REGION Network 9
   RUNG wire#powerrail
      Contact( "DB120".Static_81 )
      Contact( "TsinReq6" )
      wire#w1
      Coil( "DB127".Static_82 )
   END_RUNG
   RUNG wire#powerrail
      Contact( "DB120".Static_89 )
      Contact( "DB88".Static_8 )
   END_RUNG wire#w1
   // the same network as SCL:
   "DB127".Static_82 := ("DB120".Static_81 AND "TsinReq6") OR ("DB120".Static_89 AND "DB88".Static_8);
END_REGION

REGION Network 10
   RUNG wire#powerrail
      Contact( "DB120".Static_80 )
      I_Contact( "DB121".Static_75 )
      wire#w1
      Contact( "DB88".Static_17 )
      Coil( "DB127".Static_89 )
   END_RUNG
   RUNG wire#powerrail
      Contact( "DB120".Static_88 )
      I_Contact( "DB121".Static_75 )
   END_RUNG wire#w1
   RUNG wire#powerrail
      Contact( "DB120".Static_82 )
      I_Contact( "DB88".Static_8 )
   END_RUNG wire#w1
   // the same network as SCL:
   "DB127".Static_89 := (("DB120".Static_80 AND NOT "DB121".Static_75) OR ("DB120".Static_88 AND NOT "DB121".Static_75) OR ("DB120".Static_82 AND NOT "DB88".Static_8)) AND "DB88".Static_17;
END_REGION

REGION Network 11
   #_w1 := "DB121".Static_75 AND NOT "flReqMch6";   // rising edge
   "flReqMch6" := "DB121".Static_75;
   "DB127".Static_83 := ("DB120".Static_88 AND ("MC006-CO" OR "DB88".Static_8)) OR ("DB120".Static_84 AND NOT "DB121".Static_94 AND NOT "DB88".Static_19) OR ("DB120".Static_82 AND ("DB88".Static_19 OR "DB121".Static_94 OR "DB121".Static_75) AND "DB88".Static_8) OR (#_w1 AND "DB120".Static_82 AND "DB88".Static_8);
END_REGION

REGION Network 12
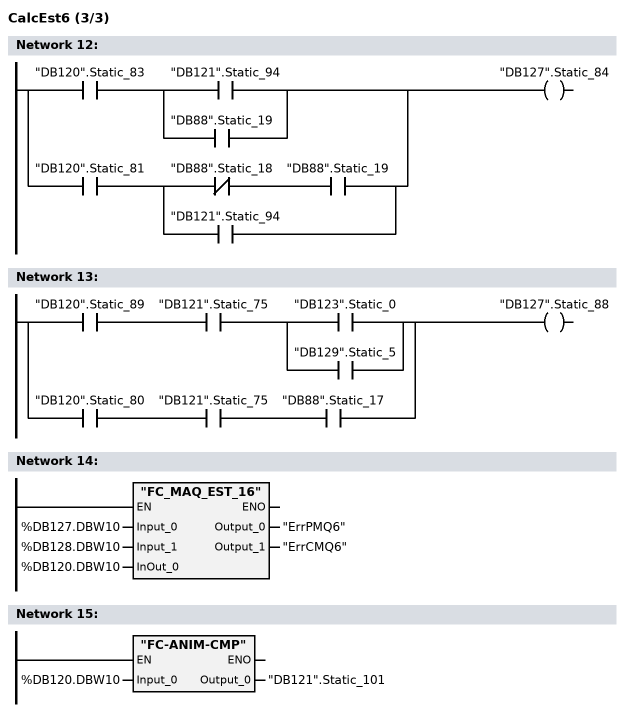
   "DB127".Static_84 := ("DB120".Static_83 AND ("DB121".Static_94 OR "DB88".Static_19)) OR ("DB120".Static_81 AND ("DB121".Static_94 OR (NOT "DB88".Static_18 AND "DB88".Static_19)));
END_REGION

REGION Network 13
   "DB127".Static_88 := ("DB120".Static_89 AND "DB121".Static_75 AND ("DB123".Static_0 OR "DB129".Static_5)) OR ("DB120".Static_80 AND "DB121".Static_75 AND "DB88".Static_17);
END_REGION

REGION Network 14
   RUNG wire#powerrail
      "FC_MAQ_EST_16"(Input_0 := %DB127.DBW10, Input_1 := %DB128.DBW10, Output_0 => "ErrPMQ6", Output_1 => "ErrCMQ6", InOut_0 := %DB120.DBW10)
   END_RUNG
   // the same network as SCL:
   "FC_MAQ_EST_16"(Input_0 := %DB127.DBW10,
                   Input_1 := %DB128.DBW10,
                   InOut_0 := %DB120.DBW10,
                   Output_0 => "ErrPMQ6",
                   Output_1 => "ErrCMQ6");
END_REGION

REGION Network 15
   RUNG wire#powerrail
      "FC-ANIM-CMP"(Input_0 := %DB120.DBW10, Output_0 => "DB121".Static_101)
   END_RUNG
   // the same network as SCL:
   "FC-ANIM-CMP"(Input_0 := %DB120.DBW10, Output_0 => "DB121".Static_101);
END_REGION
END_FUNCTION

// folder: Compresores/Baja

FUNCTION "AutoCmpBaja" : Void   // FC24, LAD
{ S7_Optimized_Access := 'FALSE' }
VERSION : 0.1
   VAR_TEMP   // added for the SCL form of the ladder/FBD networks
      _w1 : Bool;
      _s5time1 : S5Time;
      _w2 : Bool;
   END_VAR
BEGIN

REGION Network 1 (STL)
         A(;
         L     "CmpBajaAuto".Static_10;
         L     "CmpBajaAuto".Static_5;
         <=R;
         );
         JNB   M001;
         L     "CmpBajaAuto".Static_5;
         L     1;
         +R;
         T     "CmpBajaAuto".Static_10;
   M001: NOP   0;
END_REGION

REGION Network 2 (STL)
         A(;
         L     "CmpBajaAuto".Static_11;
         L     "CmpBajaAuto".Static_6;
         <=R;
         );
         JNB   M002;
         L     "CmpBajaAuto".Static_6;
         L     1;
         +R;
         T     "CmpBajaAuto".Static_11;
   M002: NOP   0;
END_REGION

REGION Network 3 (STL)
         A(;
         L     "CmpBajaAuto".Static_12;
         L     "CmpBajaAuto".Static_7;
         <=R;
         );
         JNB   M003;
         L     "CmpBajaAuto".Static_7;
         L     1;
         +R;
         T     "CmpBajaAuto".Static_12;
   M003: NOP   0;
END_REGION

REGION Network 4 (STL)
         A(;
         L     "CmpBajaAuto".Static_13;
         L     "CmpBajaAuto".Static_8;
         <=R;
         );
         JNB   M004;
         L     "CmpBajaAuto".Static_8;
         L     1;
         +R;
         T     "CmpBajaAuto".Static_13;
   M004: NOP   0;
END_REGION

REGION Network 5 (STL)
         A(;
         L     "CmpBajaAuto".Static_14;
         L     "CmpBajaAuto".Static_9;
         <=R;
         );
         JNB   M005;
         L     "CmpBajaAuto".Static_9;
         L     1;
         +R;
         T     "CmpBajaAuto".Static_14;
   M005: NOP   0;
END_REGION

REGION Network 6
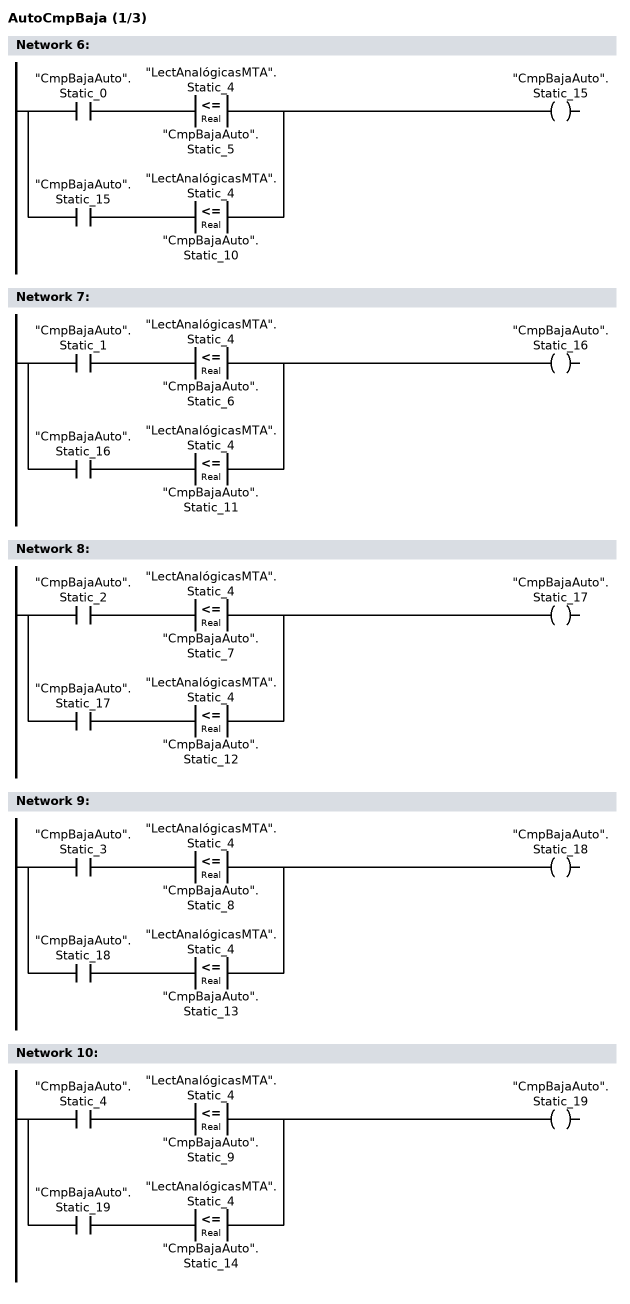
   "CmpBajaAuto".Static_15 := ("CmpBajaAuto".Static_0 AND ("LectAnalógicasMTA".Static_4 <= "CmpBajaAuto".Static_5)) OR ("CmpBajaAuto".Static_15 AND ("LectAnalógicasMTA".Static_4 <= "CmpBajaAuto".Static_10));
END_REGION

REGION Network 7
   "CmpBajaAuto".Static_16 := ("CmpBajaAuto".Static_1 AND ("LectAnalógicasMTA".Static_4 <= "CmpBajaAuto".Static_6)) OR ("CmpBajaAuto".Static_16 AND ("LectAnalógicasMTA".Static_4 <= "CmpBajaAuto".Static_11));
END_REGION

REGION Network 8
   "CmpBajaAuto".Static_17 := ("CmpBajaAuto".Static_2 AND ("LectAnalógicasMTA".Static_4 <= "CmpBajaAuto".Static_7)) OR ("CmpBajaAuto".Static_17 AND ("LectAnalógicasMTA".Static_4 <= "CmpBajaAuto".Static_12));
END_REGION

REGION Network 9
   "CmpBajaAuto".Static_18 := ("CmpBajaAuto".Static_3 AND ("LectAnalógicasMTA".Static_4 <= "CmpBajaAuto".Static_8)) OR ("CmpBajaAuto".Static_18 AND ("LectAnalógicasMTA".Static_4 <= "CmpBajaAuto".Static_13));
END_REGION

REGION Network 10
   "CmpBajaAuto".Static_19 := ("CmpBajaAuto".Static_4 AND ("LectAnalógicasMTA".Static_4 <= "CmpBajaAuto".Static_9)) OR ("CmpBajaAuto".Static_19 AND ("LectAnalógicasMTA".Static_4 <= "CmpBajaAuto".Static_14));
END_REGION

REGION Network 11
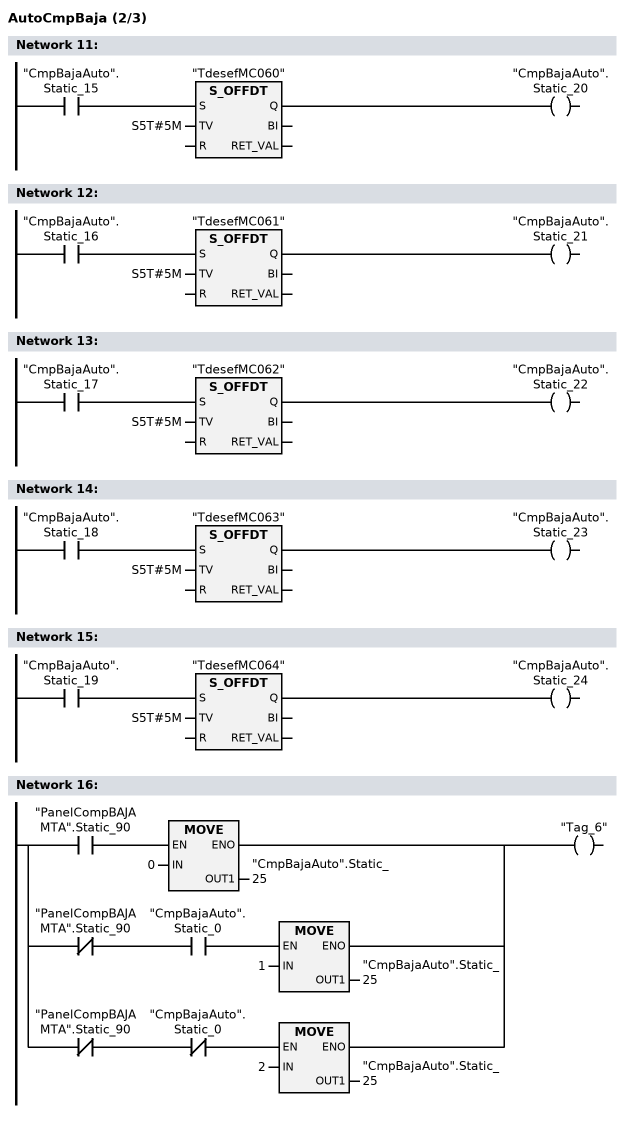
   RUNG wire#powerrail
      Contact( "CmpBajaAuto".Static_15 )
      S_OFFDT(T_NO := "TdesefMC060", TV := S5T#5M, R :=, BI =>, RET_VAL =>)
      Coil( "CmpBajaAuto".Static_20 )
   END_RUNG
   // the same network as SCL:
   #_s5time1 := S_OFFDT(T_NO := "TdesefMC060", TV := S5T#5M, S := "CmpBajaAuto".Static_15, Q => #_w1);
   "CmpBajaAuto".Static_20 := #_w1;
END_REGION

REGION Network 12
   RUNG wire#powerrail
      Contact( "CmpBajaAuto".Static_16 )
      S_OFFDT(T_NO := "TdesefMC061", TV := S5T#5M, R :=, BI =>, RET_VAL =>)
      Coil( "CmpBajaAuto".Static_21 )
   END_RUNG
   // the same network as SCL:
   #_s5time1 := S_OFFDT(T_NO := "TdesefMC061", TV := S5T#5M, S := "CmpBajaAuto".Static_16, Q => #_w1);
   "CmpBajaAuto".Static_21 := #_w1;
END_REGION

REGION Network 13
   RUNG wire#powerrail
      Contact( "CmpBajaAuto".Static_17 )
      S_OFFDT(T_NO := "TdesefMC062", TV := S5T#5M, R :=, BI =>, RET_VAL =>)
      Coil( "CmpBajaAuto".Static_22 )
   END_RUNG
   // the same network as SCL:
   #_s5time1 := S_OFFDT(T_NO := "TdesefMC062", TV := S5T#5M, S := "CmpBajaAuto".Static_17, Q => #_w1);
   "CmpBajaAuto".Static_22 := #_w1;
END_REGION

REGION Network 14
   RUNG wire#powerrail
      Contact( "CmpBajaAuto".Static_18 )
      S_OFFDT(T_NO := "TdesefMC063", TV := S5T#5M, R :=, BI =>, RET_VAL =>)
      Coil( "CmpBajaAuto".Static_23 )
   END_RUNG
   // the same network as SCL:
   #_s5time1 := S_OFFDT(T_NO := "TdesefMC063", TV := S5T#5M, S := "CmpBajaAuto".Static_18, Q => #_w1);
   "CmpBajaAuto".Static_23 := #_w1;
END_REGION

REGION Network 15
   RUNG wire#powerrail
      Contact( "CmpBajaAuto".Static_19 )
      S_OFFDT(T_NO := "TdesefMC064", TV := S5T#5M, R :=, BI =>, RET_VAL =>)
      Coil( "CmpBajaAuto".Static_24 )
   END_RUNG
   // the same network as SCL:
   #_s5time1 := S_OFFDT(T_NO := "TdesefMC064", TV := S5T#5M, S := "CmpBajaAuto".Static_19, Q => #_w1);
   "CmpBajaAuto".Static_24 := #_w1;
END_REGION

REGION Network 16
   RUNG wire#powerrail
      Contact( "PanelCompBAJA MTA".Static_90 )
      { S7_GenerateENO := "TRUE" } Move(in := 0, out1 => "CmpBajaAuto".Static_25)
      wire#w1
      Coil( "Tag_6" )
   END_RUNG
   RUNG wire#powerrail
      I_Contact( "PanelCompBAJA MTA".Static_90 )
      Contact( "CmpBajaAuto".Static_0 )
      { S7_GenerateENO := "TRUE" } Move(in := 1, out1 => "CmpBajaAuto".Static_25)
   END_RUNG wire#w1
   RUNG wire#powerrail
      I_Contact( "PanelCompBAJA MTA".Static_90 )
      I_Contact( "CmpBajaAuto".Static_0 )
      { S7_GenerateENO := "TRUE" } Move(in := 2, out1 => "CmpBajaAuto".Static_25)
   END_RUNG wire#w1
   // the same network as SCL:
   // ENO of a box is taken as its EN; it also drops when the box reports an error
   IF "PanelCompBAJA MTA".Static_90 THEN "CmpBajaAuto".Static_25 := 0; END_IF;
   #_w1 := NOT "PanelCompBAJA MTA".Static_90 AND "CmpBajaAuto".Static_0;
   IF #_w1 THEN "CmpBajaAuto".Static_25 := 1; END_IF;
   #_w2 := NOT "PanelCompBAJA MTA".Static_90 AND NOT "CmpBajaAuto".Static_0;
   IF #_w2 THEN "CmpBajaAuto".Static_25 := 2; END_IF;
   "Tag_6" := "PanelCompBAJA MTA".Static_90 OR #_w1 OR #_w2;
END_REGION

REGION Network 17
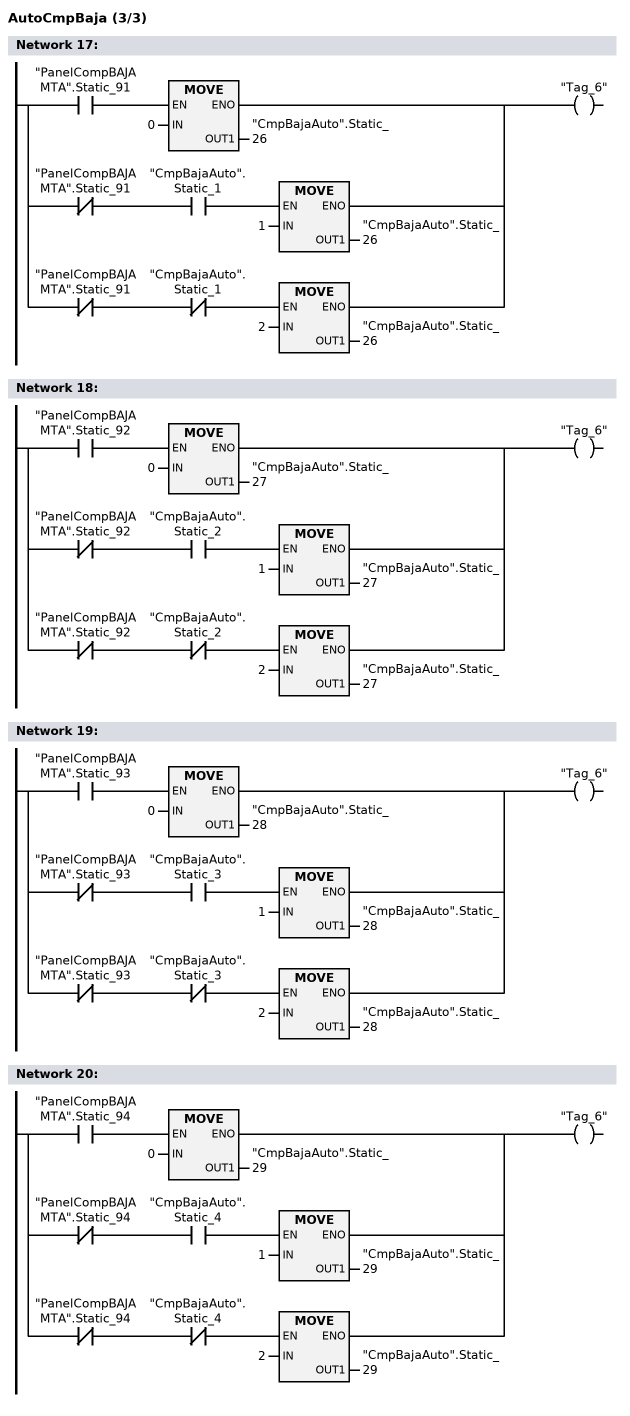
   RUNG wire#powerrail
      Contact( "PanelCompBAJA MTA".Static_91 )
      { S7_GenerateENO := "TRUE" } Move(in := 0, out1 => "CmpBajaAuto".Static_26)
      wire#w1
      Coil( "Tag_6" )
   END_RUNG
   RUNG wire#powerrail
      I_Contact( "PanelCompBAJA MTA".Static_91 )
      Contact( "CmpBajaAuto".Static_1 )
      { S7_GenerateENO := "TRUE" } Move(in := 1, out1 => "CmpBajaAuto".Static_26)
   END_RUNG wire#w1
   RUNG wire#powerrail
      I_Contact( "PanelCompBAJA MTA".Static_91 )
      I_Contact( "CmpBajaAuto".Static_1 )
      { S7_GenerateENO := "TRUE" } Move(in := 2, out1 => "CmpBajaAuto".Static_26)
   END_RUNG wire#w1
   // the same network as SCL:
   // ENO of a box is taken as its EN; it also drops when the box reports an error
   IF "PanelCompBAJA MTA".Static_91 THEN "CmpBajaAuto".Static_26 := 0; END_IF;
   #_w1 := NOT "PanelCompBAJA MTA".Static_91 AND "CmpBajaAuto".Static_1;
   IF #_w1 THEN "CmpBajaAuto".Static_26 := 1; END_IF;
   #_w2 := NOT "PanelCompBAJA MTA".Static_91 AND NOT "CmpBajaAuto".Static_1;
   IF #_w2 THEN "CmpBajaAuto".Static_26 := 2; END_IF;
   "Tag_6" := "PanelCompBAJA MTA".Static_91 OR #_w1 OR #_w2;
END_REGION

REGION Network 18
   RUNG wire#powerrail
      Contact( "PanelCompBAJA MTA".Static_92 )
      { S7_GenerateENO := "TRUE" } Move(in := 0, out1 => "CmpBajaAuto".Static_27)
      wire#w1
      Coil( "Tag_6" )
   END_RUNG
   RUNG wire#powerrail
      I_Contact( "PanelCompBAJA MTA".Static_92 )
      Contact( "CmpBajaAuto".Static_2 )
      { S7_GenerateENO := "TRUE" } Move(in := 1, out1 => "CmpBajaAuto".Static_27)
   END_RUNG wire#w1
   RUNG wire#powerrail
      I_Contact( "PanelCompBAJA MTA".Static_92 )
      I_Contact( "CmpBajaAuto".Static_2 )
      { S7_GenerateENO := "TRUE" } Move(in := 2, out1 => "CmpBajaAuto".Static_27)
   END_RUNG wire#w1
   // the same network as SCL:
   // ENO of a box is taken as its EN; it also drops when the box reports an error
   IF "PanelCompBAJA MTA".Static_92 THEN "CmpBajaAuto".Static_27 := 0; END_IF;
   #_w1 := NOT "PanelCompBAJA MTA".Static_92 AND "CmpBajaAuto".Static_2;
   IF #_w1 THEN "CmpBajaAuto".Static_27 := 1; END_IF;
   #_w2 := NOT "PanelCompBAJA MTA".Static_92 AND NOT "CmpBajaAuto".Static_2;
   IF #_w2 THEN "CmpBajaAuto".Static_27 := 2; END_IF;
   "Tag_6" := "PanelCompBAJA MTA".Static_92 OR #_w1 OR #_w2;
END_REGION

REGION Network 19
   RUNG wire#powerrail
      Contact( "PanelCompBAJA MTA".Static_93 )
      { S7_GenerateENO := "TRUE" } Move(in := 0, out1 => "CmpBajaAuto".Static_28)
      wire#w1
      Coil( "Tag_6" )
   END_RUNG
   RUNG wire#powerrail
      I_Contact( "PanelCompBAJA MTA".Static_93 )
      Contact( "CmpBajaAuto".Static_3 )
      { S7_GenerateENO := "TRUE" } Move(in := 1, out1 => "CmpBajaAuto".Static_28)
   END_RUNG wire#w1
   RUNG wire#powerrail
      I_Contact( "PanelCompBAJA MTA".Static_93 )
      I_Contact( "CmpBajaAuto".Static_3 )
      { S7_GenerateENO := "TRUE" } Move(in := 2, out1 => "CmpBajaAuto".Static_28)
   END_RUNG wire#w1
   // the same network as SCL:
   // ENO of a box is taken as its EN; it also drops when the box reports an error
   IF "PanelCompBAJA MTA".Static_93 THEN "CmpBajaAuto".Static_28 := 0; END_IF;
   #_w1 := NOT "PanelCompBAJA MTA".Static_93 AND "CmpBajaAuto".Static_3;
   IF #_w1 THEN "CmpBajaAuto".Static_28 := 1; END_IF;
   #_w2 := NOT "PanelCompBAJA MTA".Static_93 AND NOT "CmpBajaAuto".Static_3;
   IF #_w2 THEN "CmpBajaAuto".Static_28 := 2; END_IF;
   "Tag_6" := "PanelCompBAJA MTA".Static_93 OR #_w1 OR #_w2;
END_REGION

REGION Network 20
   RUNG wire#powerrail
      Contact( "PanelCompBAJA MTA".Static_94 )
      { S7_GenerateENO := "TRUE" } Move(in := 0, out1 => "CmpBajaAuto".Static_29)
      wire#w1
      Coil( "Tag_6" )
   END_RUNG
   RUNG wire#powerrail
      I_Contact( "PanelCompBAJA MTA".Static_94 )
      Contact( "CmpBajaAuto".Static_4 )
      { S7_GenerateENO := "TRUE" } Move(in := 1, out1 => "CmpBajaAuto".Static_29)
   END_RUNG wire#w1
   RUNG wire#powerrail
      I_Contact( "PanelCompBAJA MTA".Static_94 )
      I_Contact( "CmpBajaAuto".Static_4 )
      { S7_GenerateENO := "TRUE" } Move(in := 2, out1 => "CmpBajaAuto".Static_29)
   END_RUNG wire#w1
   // the same network as SCL:
   // ENO of a box is taken as its EN; it also drops when the box reports an error
   IF "PanelCompBAJA MTA".Static_94 THEN "CmpBajaAuto".Static_29 := 0; END_IF;
   #_w1 := NOT "PanelCompBAJA MTA".Static_94 AND "CmpBajaAuto".Static_4;
   IF #_w1 THEN "CmpBajaAuto".Static_29 := 1; END_IF;
   #_w2 := NOT "PanelCompBAJA MTA".Static_94 AND NOT "CmpBajaAuto".Static_4;
   IF #_w2 THEN "CmpBajaAuto".Static_29 := 2; END_IF;
   "Tag_6" := "PanelCompBAJA MTA".Static_94 OR #_w1 OR #_w2;
END_REGION
END_FUNCTION

// folder: Entradas analógicas

FUNCTION "LecturasAnalógicasMTA" : Void   // FC15, LAD
{ S7_Optimized_Access := 'FALSE' }
VERSION : 0.1
BEGIN

REGION Network 1
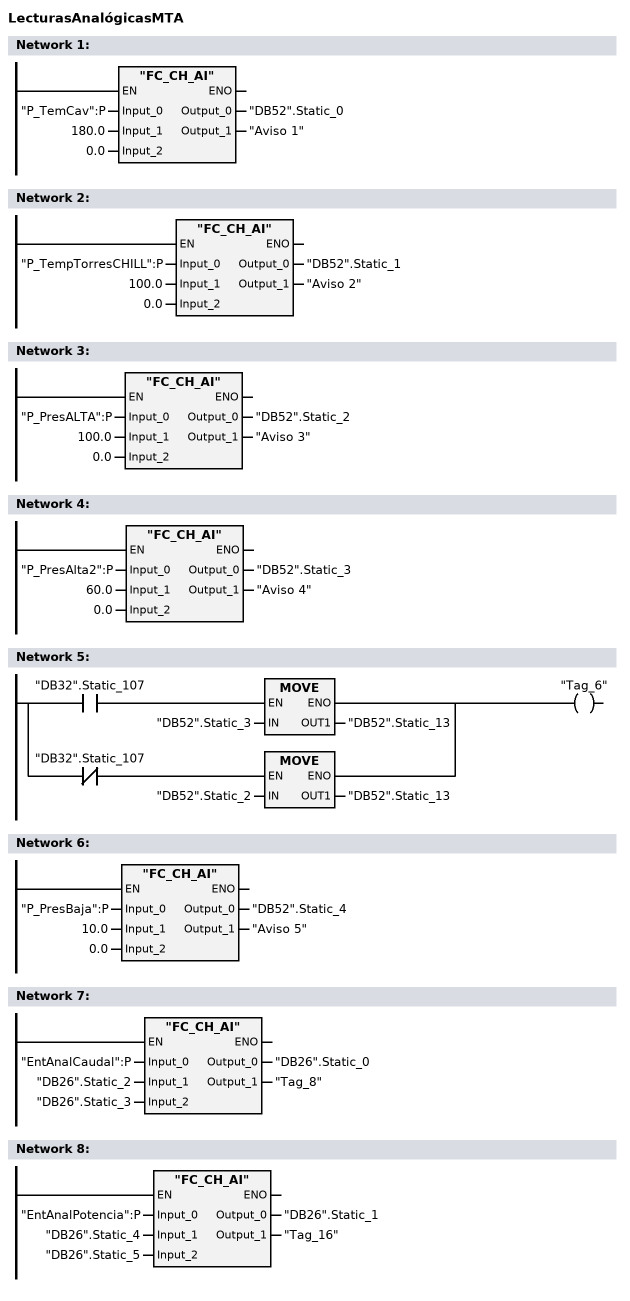
   RUNG wire#powerrail
      "FC_CH_AI"(Input_0 := "P_TemCav":P, Input_1 := 180.0, Input_2 := 0.0, Output_0 => "DB52".Static_0, Output_1 => "Aviso 1")
   END_RUNG
   // the same network as SCL:
   "FC_CH_AI"(Input_0 := "P_TemCav":P,
              Input_1 := 180.0,
              Input_2 := 0.0,
              Output_0 => "DB52".Static_0,
              Output_1 => "Aviso 1");
END_REGION

REGION Network 2
   RUNG wire#powerrail
      "FC_CH_AI"(Input_0 := "P_TempTorresCHILL":P, Input_1 := 100.0, Input_2 := 0.0, Output_0 => "DB52".Static_1, Output_1 => "Aviso 2")
   END_RUNG
   // the same network as SCL:
   "FC_CH_AI"(Input_0 := "P_TempTorresCHILL":P,
              Input_1 := 100.0,
              Input_2 := 0.0,
              Output_0 => "DB52".Static_1,
              Output_1 => "Aviso 2");
END_REGION

REGION Network 3
   RUNG wire#powerrail
      "FC_CH_AI"(Input_0 := "P_PresALTA":P, Input_1 := 100.0, Input_2 := 0.0, Output_0 => "DB52".Static_2, Output_1 => "Aviso 3")
   END_RUNG
   // the same network as SCL:
   "FC_CH_AI"(Input_0 := "P_PresALTA":P,
              Input_1 := 100.0,
              Input_2 := 0.0,
              Output_0 => "DB52".Static_2,
              Output_1 => "Aviso 3");
END_REGION

REGION Network 4
   RUNG wire#powerrail
      "FC_CH_AI"(Input_0 := "P_PresAlta2":P, Input_1 := 60.0, Input_2 := 0.0, Output_0 => "DB52".Static_3, Output_1 => "Aviso 4")
   END_RUNG
   // the same network as SCL:
   "FC_CH_AI"(Input_0 := "P_PresAlta2":P,
              Input_1 := 60.0,
              Input_2 := 0.0,
              Output_0 => "DB52".Static_3,
              Output_1 => "Aviso 4");
END_REGION

REGION Network 5
   RUNG wire#powerrail
      Contact( "DB32".Static_107 )
      { S7_GenerateENO := "TRUE" } Move(in := "DB52".Static_3, out1 => "DB52".Static_13)
      wire#w1
      Coil( "Tag_6" )
   END_RUNG
   RUNG wire#powerrail
      I_Contact( "DB32".Static_107 )
      { S7_GenerateENO := "TRUE" } Move(in := "DB52".Static_2, out1 => "DB52".Static_13)
   END_RUNG wire#w1
   // the same network as SCL:
   // ENO of a box is taken as its EN; it also drops when the box reports an error
   IF "DB32".Static_107 THEN "DB52".Static_13 := "DB52".Static_3; END_IF;
   IF NOT "DB32".Static_107 THEN "DB52".Static_13 := "DB52".Static_2; END_IF;
   "Tag_6" := "DB32".Static_107 OR NOT "DB32".Static_107;
END_REGION

REGION Network 6
   RUNG wire#powerrail
      "FC_CH_AI"(Input_0 := "P_PresBaja":P, Input_1 := 10.0, Input_2 := 0.0, Output_0 => "DB52".Static_4, Output_1 => "Aviso 5")
   END_RUNG
   // the same network as SCL:
   "FC_CH_AI"(Input_0 := "P_PresBaja":P,
              Input_1 := 10.0,
              Input_2 := 0.0,
              Output_0 => "DB52".Static_4,
              Output_1 => "Aviso 5");
END_REGION

REGION Network 7
   RUNG wire#powerrail
      "FC_CH_AI"(Input_0 := "EntAnalCaudal":P, Input_1 := "DB26".Static_2, Input_2 := "DB26".Static_3, Output_0 => "DB26".Static_0, Output_1 => "Tag_8")
   END_RUNG
   // the same network as SCL:
   "FC_CH_AI"(Input_0 := "EntAnalCaudal":P,
              Input_1 := "DB26".Static_2,
              Input_2 := "DB26".Static_3,
              Output_0 => "DB26".Static_0,
              Output_1 => "Tag_8");
END_REGION

REGION Network 8
   RUNG wire#powerrail
      "FC_CH_AI"(Input_0 := "EntAnalPotencia":P, Input_1 := "DB26".Static_4, Input_2 := "DB26".Static_5, Output_0 => "DB26".Static_1, Output_1 => "Tag_16")
   END_RUNG
   // the same network as SCL:
   "FC_CH_AI"(Input_0 := "EntAnalPotencia":P,
              Input_1 := "DB26".Static_4,
              Input_2 := "DB26".Static_5,
              Output_0 => "DB26".Static_1,
              Output_1 => "Tag_16");
END_REGION
END_FUNCTION

// folder: Horas de Marcha

ORGANIZATION_BLOCK "CYC_INT5"   // OB35, LAD
{ S7_Optimized_Access := 'FALSE' }
VERSION : 0.1
   VAR_TEMP   // added for the SCL form of the ladder/FBD networks
      _w1 : Bool;
      _w2 : Bool;
      _w3 : Bool;
      _w4 : Bool;
   END_VAR
BEGIN

REGION Network 1 (STL)
         A     "MC001";
         A     "MC001-CO";
         =     <??.?>;
         A     <??.?>;
         A(;
         L     "DB73".Static_27;
         L     600;
         <I;
         );
         JNB   M001;
         L     1;
         L     "DB73".Static_27;
         +D;
         T     "DB73".Static_27;
   M001: NOP   0;
         A     <??.?>;
         A(;
         L     "DB73".Static_27;
         L     600;
         >=I;
         );
         =     <??.?>;
         A     <??.?>;
         JNB   M002;
         L     1;
         L     "DB73".Static_6;
         +D;
         T     "DB73".Static_6;
   M002: NOP   0;
         A     <??.?>;
         JNB   M003;
         L     0;
         T     "DB73".Static_27;
   M003: NOP   0;
         A     <??.?>;
         A(;
         L     "DB73".Static_6;
         L     60;
         >=I;
         );
         =     <??.?>;
         A     <??.?>;
         JNB   M004;
         L     1;
         L     "DB73".Static_0;
         +D;
         T     "DB73".Static_0;
   M004: NOP   0;
         A     <??.?>;
         JNB   M005;
         L     0;
         T     "DB73".Static_6;
   M005: NOP   0;
END_REGION

REGION Network 2 (STL)
         A     "MC002";
         A     "MC002-CO";
         =     <??.?>;
         A     <??.?>;
         A(;
         L     "DB73".Static_28;
         L     600;
         <I;
         );
         JNB   M006;
         L     1;
         L     "DB73".Static_28;
         +D;
         T     "DB73".Static_28;
   M006: NOP   0;
         A     <??.?>;
         A(;
         L     "DB73".Static_28;
         L     600;
         >=I;
         );
         =     <??.?>;
         A     <??.?>;
         JNB   M007;
         L     1;
         L     "DB73".Static_7;
         +D;
         T     "DB73".Static_7;
   M007: NOP   0;
         A     <??.?>;
         JNB   M008;
         L     0;
         T     "DB73".Static_28;
   M008: NOP   0;
         A     <??.?>;
         A(;
         L     "DB73".Static_7;
         L     60;
         >=I;
         );
         =     <??.?>;
         A     <??.?>;
         JNB   M009;
         L     1;
         L     "DB73".Static_1;
         +D;
         T     "DB73".Static_1;
   M009: NOP   0;
         A     <??.?>;
         JNB   M010;
         L     0;
         T     "DB73".Static_7;
   M010: NOP   0;
END_REGION

REGION Network 3 (STL)
         A     "MC003";
         A     "MC003-CO";
         =     <??.?>;
         A     <??.?>;
         A(;
         L     "DB73".Static_29;
         L     600;
         <I;
         );
         JNB   M011;
         L     1;
         L     "DB73".Static_29;
         +D;
         T     "DB73".Static_29;
   M011: NOP   0;
         A     <??.?>;
         A(;
         L     "DB73".Static_29;
         L     600;
         >=I;
         );
         =     <??.?>;
         A     <??.?>;
         JNB   M012;
         L     1;
         L     "DB73".Static_8;
         +D;
         T     "DB73".Static_8;
   M012: NOP   0;
         A     <??.?>;
         JNB   M013;
         L     0;
         T     "DB73".Static_29;
   M013: NOP   0;
         A     <??.?>;
         A(;
         L     "DB73".Static_8;
         L     60;
         >=I;
         );
         =     <??.?>;
         A     <??.?>;
         JNB   M014;
         L     1;
         L     "DB73".Static_2;
         +D;
         T     "DB73".Static_2;
   M014: NOP   0;
         A     <??.?>;
         JNB   M015;
         L     0;
         T     "DB73".Static_8;
   M015: NOP   0;
END_REGION

REGION Network 4 (STL)
         A     "MC004";
         A     "MC004-CO";
         =     <??.?>;
         A     <??.?>;
         A(;
         L     "DB73".Static_30;
         L     600;
         <I;
         );
         JNB   M016;
         L     1;
         L     "DB73".Static_30;
         +D;
         T     "DB73".Static_30;
   M016: NOP   0;
         A     <??.?>;
         A(;
         L     "DB73".Static_30;
         L     600;
         >=I;
         );
         =     <??.?>;
         A     <??.?>;
         JNB   M017;
         L     1;
         L     "DB73".Static_9;
         +D;
         T     "DB73".Static_9;
   M017: NOP   0;
         A     <??.?>;
         JNB   M018;
         L     0;
         T     "DB73".Static_30;
   M018: NOP   0;
         A     <??.?>;
         A(;
         L     "DB73".Static_9;
         L     60;
         >=I;
         );
         =     <??.?>;
         A     <??.?>;
         JNB   M019;
         L     1;
         L     "DB73".Static_3;
         +D;
         T     "DB73".Static_3;
   M019: NOP   0;
         A     <??.?>;
         JNB   M020;
         L     0;
         T     "DB73".Static_9;
   M020: NOP   0;
END_REGION

REGION Network 5 (STL)
         A     "MC005";
         A     "MC005-CO";
         =     <??.?>;
         A     <??.?>;
         A(;
         L     "DB73".Static_31;
         L     600;
         <I;
         );
         JNB   M021;
         L     1;
         L     "DB73".Static_31;
         +D;
         T     "DB73".Static_31;
   M021: NOP   0;
         A     <??.?>;
         A(;
         L     "DB73".Static_31;
         L     600;
         >=I;
         );
         =     <??.?>;
         A     <??.?>;
         JNB   M022;
         L     1;
         L     "DB73".Static_10;
         +D;
         T     "DB73".Static_10;
   M022: NOP   0;
         A     <??.?>;
         JNB   M023;
         L     0;
         T     "DB73".Static_31;
   M023: NOP   0;
         A     <??.?>;
         A(;
         L     "DB73".Static_10;
         L     60;
         >=I;
         );
         =     <??.?>;
         A     <??.?>;
         JNB   M024;
         L     1;
         L     "DB73".Static_4;
         +D;
         T     "DB73".Static_4;
   M024: NOP   0;
         A     <??.?>;
         JNB   M025;
         L     0;
         T     "DB73".Static_10;
   M025: NOP   0;
END_REGION

REGION Network 6 (STL)
         A     "MC006";
         A     "MC006-CO";
         =     <??.?>;
         A     <??.?>;
         A(;
         L     "DB73".Static_32;
         L     600;
         <I;
         );
         JNB   M026;
         L     1;
         L     "DB73".Static_32;
         +D;
         T     "DB73".Static_32;
   M026: NOP   0;
         A     <??.?>;
         A(;
         L     "DB73".Static_32;
         L     600;
         >=I;
         );
         =     <??.?>;
         A     <??.?>;
         JNB   M027;
         L     1;
         L     "DB73".Static_11;
         +D;
         T     "DB73".Static_11;
   M027: NOP   0;
         A     <??.?>;
         JNB   M028;
         L     0;
         T     "DB73".Static_32;
   M028: NOP   0;
         A     <??.?>;
         A(;
         L     "DB73".Static_11;
         L     60;
         >=I;
         );
         =     <??.?>;
         A     <??.?>;
         JNB   M029;
         L     1;
         L     "DB73".Static_5;
         +D;
         T     "DB73".Static_5;
   M029: NOP   0;
         A     <??.?>;
         JNB   M030;
         L     0;
         T     "DB73".Static_11;
   M030: NOP   0;
END_REGION

REGION Network 7
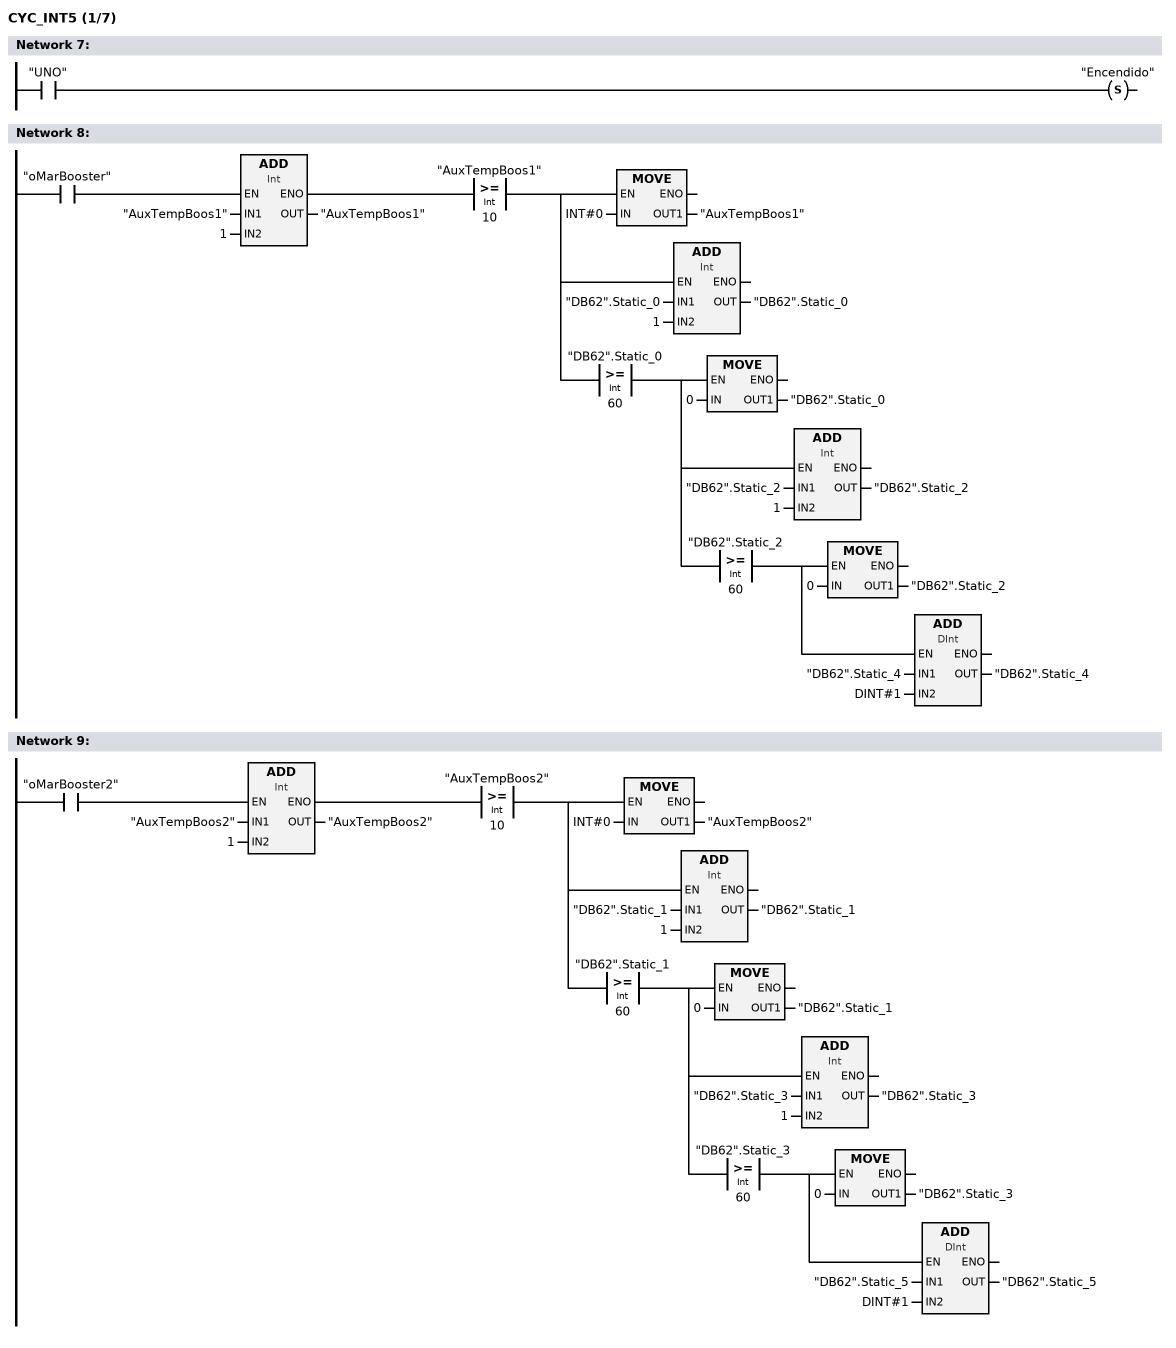
   RUNG wire#powerrail
      Contact( "UNO" )
      S_Coil( "Encendido" )
   END_RUNG
   // the same network as SCL:
   IF "UNO" THEN "Encendido" := TRUE; END_IF;
END_REGION

REGION Network 8
   RUNG wire#powerrail
      Contact( "oMarBooster" )
      { S7_Templates := "SrcType := Int"; S7_GenerateENO := "TRUE" } Add(in1 := "AuxTempBoos1", in2 := 1, out => "AuxTempBoos1")
      { S7_Templates := "SrcType := Int" } GE_Contact(in1 := "AuxTempBoos1", in2 := 10)
      wire#w1
      { S7_GenerateENO := "TRUE" } Move(in := INT#0, out1 => "AuxTempBoos1")
   END_RUNG
   RUNG wire#w1
      { S7_Templates := "SrcType := Int"; S7_GenerateENO := "TRUE" } Add(in1 := "DB62".Static_0, in2 := 1, out => "DB62".Static_0)
   END_RUNG
   RUNG wire#w1
      { S7_Templates := "SrcType := Int" } GE_Contact(in1 := "DB62".Static_0, in2 := 60)
      wire#w2
      { S7_GenerateENO := "TRUE" } Move(in := 0, out1 => "DB62".Static_0)
   END_RUNG
   RUNG wire#w2
      { S7_Templates := "SrcType := Int"; S7_GenerateENO := "TRUE" } Add(in1 := "DB62".Static_2, in2 := 1, out => "DB62".Static_2)
   END_RUNG
   RUNG wire#w2
      { S7_Templates := "SrcType := Int" } GE_Contact(in1 := "DB62".Static_2, in2 := 60)
      wire#w3
      { S7_GenerateENO := "TRUE" } Move(in := 0, out1 => "DB62".Static_2)
   END_RUNG
   RUNG wire#w3
      { S7_Templates := "SrcType := DInt"; S7_GenerateENO := "TRUE" } Add(in1 := "DB62".Static_4, in2 := DINT#1, out => "DB62".Static_4)
   END_RUNG
   // the same network as SCL:
   // ENO of a box is taken as its EN; it also drops when the box reports an error
   IF "oMarBooster" THEN "AuxTempBoos1" := "AuxTempBoos1" + 1; END_IF;
   #_w1 := "oMarBooster" AND ("AuxTempBoos1" >= 10);
   IF #_w1 THEN
       "AuxTempBoos1" := INT#0;
       "DB62".Static_0 := "DB62".Static_0 + 1;
   END_IF;
   #_w2 := #_w1 AND ("DB62".Static_0 >= 60);
   IF #_w2 THEN
       "DB62".Static_0 := 0;
       "DB62".Static_2 := "DB62".Static_2 + 1;
   END_IF;
   #_w3 := #_w2 AND ("DB62".Static_2 >= 60);
   IF #_w3 THEN
       "DB62".Static_2 := 0;
       "DB62".Static_4 := "DB62".Static_4 + DINT#1;
   END_IF;
END_REGION

REGION Network 9
   RUNG wire#powerrail
      Contact( "oMarBooster2" )
      { S7_Templates := "SrcType := Int"; S7_GenerateENO := "TRUE" } Add(in1 := "AuxTempBoos2", in2 := 1, out => "AuxTempBoos2")
      { S7_Templates := "SrcType := Int" } GE_Contact(in1 := "AuxTempBoos2", in2 := 10)
      wire#w1
      { S7_GenerateENO := "TRUE" } Move(in := INT#0, out1 => "AuxTempBoos2")
   END_RUNG
   RUNG wire#w1
      { S7_Templates := "SrcType := Int"; S7_GenerateENO := "TRUE" } Add(in1 := "DB62".Static_1, in2 := 1, out => "DB62".Static_1)
   END_RUNG
   RUNG wire#w1
      { S7_Templates := "SrcType := Int" } GE_Contact(in1 := "DB62".Static_1, in2 := 60)
      wire#w2
      { S7_GenerateENO := "TRUE" } Move(in := 0, out1 => "DB62".Static_1)
   END_RUNG
   RUNG wire#w2
      { S7_Templates := "SrcType := Int"; S7_GenerateENO := "TRUE" } Add(in1 := "DB62".Static_3, in2 := 1, out => "DB62".Static_3)
   END_RUNG
   RUNG wire#w2
      { S7_Templates := "SrcType := Int" } GE_Contact(in1 := "DB62".Static_3, in2 := 60)
      wire#w3
      { S7_GenerateENO := "TRUE" } Move(in := 0, out1 => "DB62".Static_3)
   END_RUNG
   RUNG wire#w3
      { S7_Templates := "SrcType := DInt"; S7_GenerateENO := "TRUE" } Add(in1 := "DB62".Static_5, in2 := DINT#1, out => "DB62".Static_5)
   END_RUNG
   // the same network as SCL:
   // ENO of a box is taken as its EN; it also drops when the box reports an error
   IF "oMarBooster2" THEN "AuxTempBoos2" := "AuxTempBoos2" + 1; END_IF;
   #_w1 := "oMarBooster2" AND ("AuxTempBoos2" >= 10);
   IF #_w1 THEN
       "AuxTempBoos2" := INT#0;
       "DB62".Static_1 := "DB62".Static_1 + 1;
   END_IF;
   #_w2 := #_w1 AND ("DB62".Static_1 >= 60);
   IF #_w2 THEN
       "DB62".Static_1 := 0;
       "DB62".Static_3 := "DB62".Static_3 + 1;
   END_IF;
   #_w3 := #_w2 AND ("DB62".Static_3 >= 60);
   IF #_w3 THEN
       "DB62".Static_3 := 0;
       "DB62".Static_5 := "DB62".Static_5 + DINT#1;
   END_IF;
END_REGION

REGION Network 10